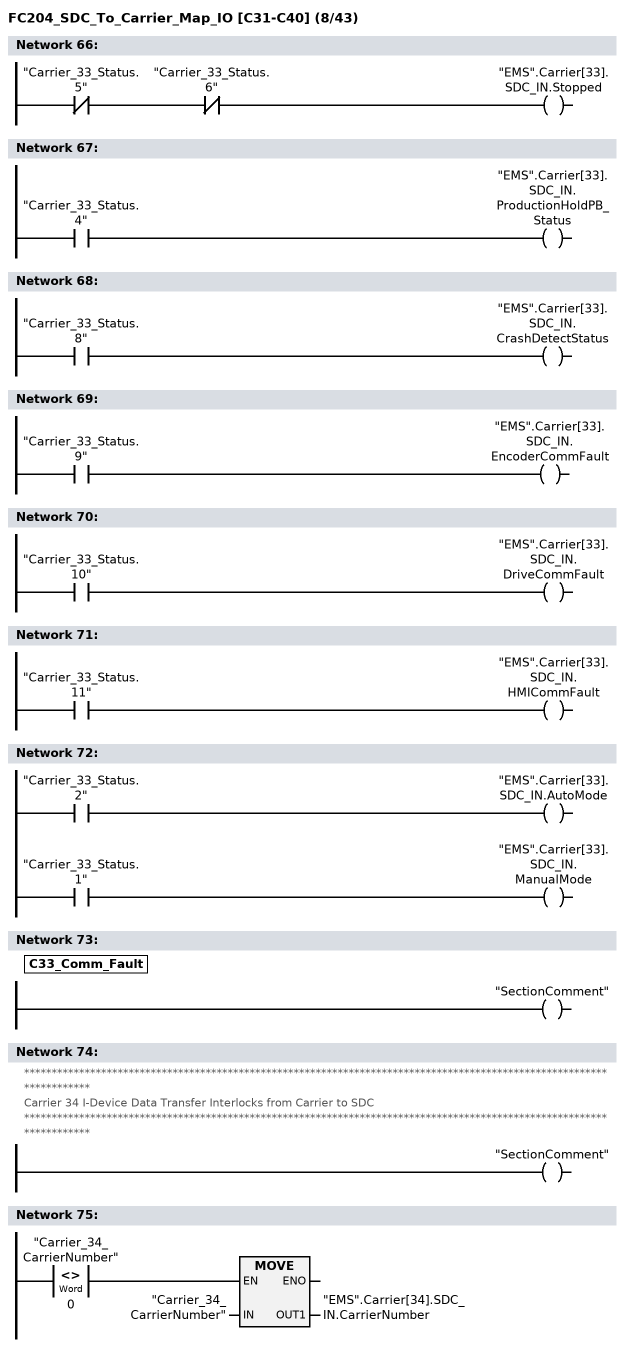
   RUNG wire#powerrail
      I_Contact( "Carrier_33_Status.5" )
      I_Contact( "Carrier_33_Status.6" )
      Coil( "EMS".Carrier[33].SDC_IN.Stopped )
   END_RUNG
   // the same network as SCL:
   "EMS".Carrier[33].SDC_IN.Stopped := NOT "Carrier_33_Status.5" AND NOT "Carrier_33_Status.6";
END_REGION

REGION Network 67
   RUNG wire#powerrail
      Contact( "Carrier_33_Status.4" )
      Coil( "EMS".Carrier[33].SDC_IN.ProductionHoldPB_Status )
   END_RUNG
   // the same network as SCL:
   "EMS".Carrier[33].SDC_IN.ProductionHoldPB_Status := "Carrier_33_Status.4";
END_REGION

REGION Network 68
   RUNG wire#powerrail
      Contact( "Carrier_33_Status.8" )
      Coil( "EMS".Carrier[33].SDC_IN.CrashDetectStatus )
   END_RUNG
   // the same network as SCL:
   "EMS".Carrier[33].SDC_IN.CrashDetectStatus := "Carrier_33_Status.8";
END_REGION

REGION Network 69
   RUNG wire#powerrail
      Contact( "Carrier_33_Status.9" )
      Coil( "EMS".Carrier[33].SDC_IN.EncoderCommFault )
   END_RUNG
   // the same network as SCL:
   "EMS".Carrier[33].SDC_IN.EncoderCommFault := "Carrier_33_Status.9";
END_REGION

REGION Network 70
   RUNG wire#powerrail
      Contact( "Carrier_33_Status.10" )
      Coil( "EMS".Carrier[33].SDC_IN.DriveCommFault )
   END_RUNG
   // the same network as SCL:
   "EMS".Carrier[33].SDC_IN.DriveCommFault := "Carrier_33_Status.10";
END_REGION

REGION Network 71
   RUNG wire#powerrail
      Contact( "Carrier_33_Status.11" )
      Coil( "EMS".Carrier[33].SDC_IN.HMICommFault )
   END_RUNG
   // the same network as SCL:
   "EMS".Carrier[33].SDC_IN.HMICommFault := "Carrier_33_Status.11";
END_REGION

REGION Network 72
   RUNG wire#powerrail
      Contact( "Carrier_33_Status.2" )
      Coil( "EMS".Carrier[33].SDC_IN.AutoMode )
   END_RUNG
   RUNG wire#powerrail
      Contact( "Carrier_33_Status.1" )
      Coil( "EMS".Carrier[33].SDC_IN.ManualMode )
   END_RUNG
   // the same network as SCL:
   "EMS".Carrier[33].SDC_IN.AutoMode := "Carrier_33_Status.2";
   "EMS".Carrier[33].SDC_IN.ManualMode := "Carrier_33_Status.1";
END_REGION

REGION Network 73
   Label( C33_Comm_Fault )
   RUNG wire#powerrail
      Coil( "SectionComment" )
   END_RUNG
   // the same network as SCL:
   C33_Comm_Fault:
   "SectionComment" := TRUE;
END_REGION

REGION Network 74
   // **********************************************************************************************************************
   // 
   // Carrier 34 I-Device Data Transfer Interlocks from Carrier to SDC
   // 
   // **********************************************************************************************************************
   RUNG wire#powerrail
      Coil( "SectionComment" )
   END_RUNG
   // the same network as SCL:
   "SectionComment" := TRUE;
END_REGION

REGION Network 75
   RUNG wire#powerrail
      { S7_Templates := "SrcType := Word" } NE_Contact(in1 := "Carrier_34_CarrierNumber", in2 := 0)
      Move(in := "Carrier_34_CarrierNumber", out1 => "EMS".Carrier[34].SDC_IN.CarrierNumber)
   END_RUNG
   // the same network as SCL:
   IF "Carrier_34_CarrierNumber" <> 0 THEN
       "EMS".Carrier[34].SDC_IN.CarrierNumber := "Carrier_34_CarrierNumber";
   END_IF;
END_REGION

REGION Network 76
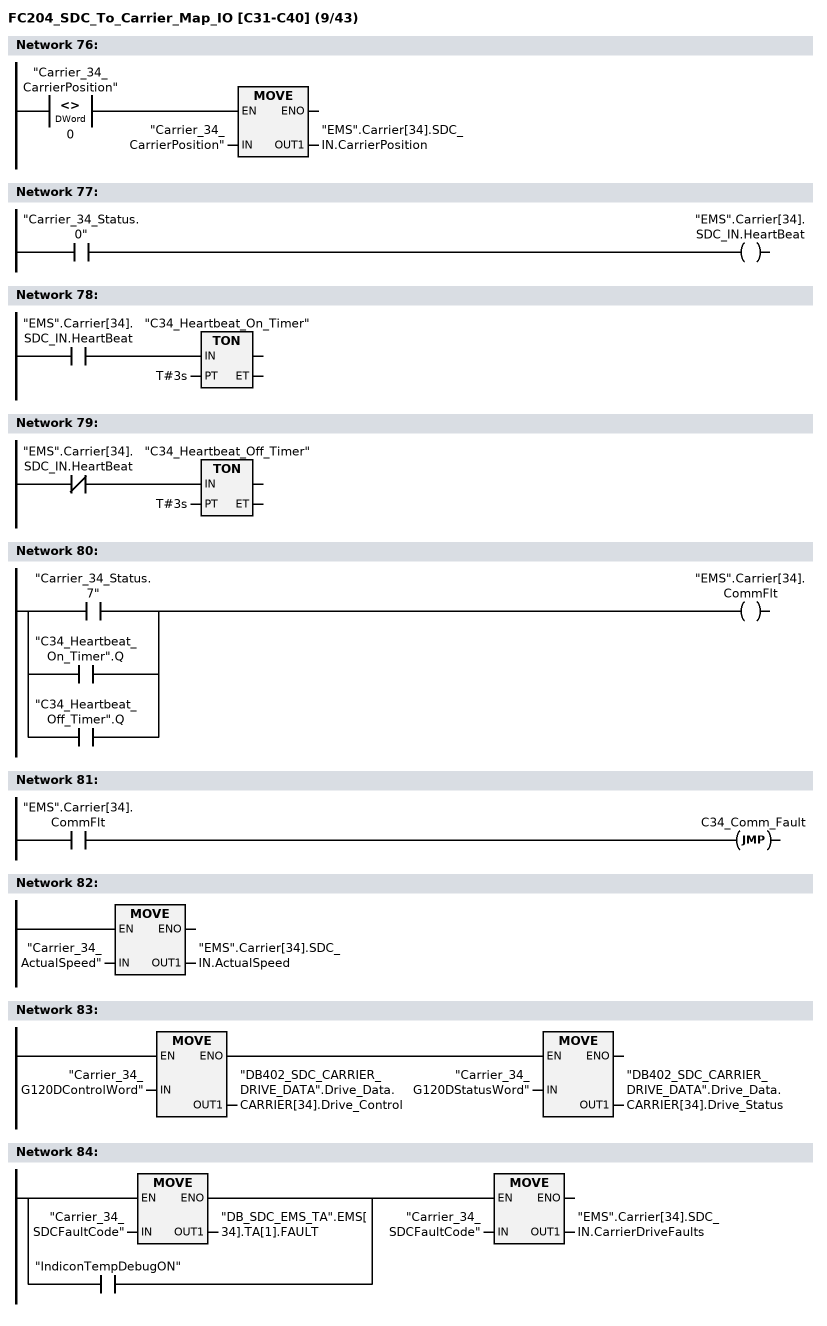
   RUNG wire#powerrail
      { S7_Templates := "SrcType := DWord" } NE_Contact(in1 := "Carrier_34_CarrierPosition", in2 := 0)
      Move(in := "Carrier_34_CarrierPosition", out1 => "EMS".Carrier[34].SDC_IN.CarrierPosition)
   END_RUNG
   // the same network as SCL:
   IF "Carrier_34_CarrierPosition" <> 0 THEN
       "EMS".Carrier[34].SDC_IN.CarrierPosition := "Carrier_34_CarrierPosition";
   END_IF;
END_REGION

REGION Network 77
   RUNG wire#powerrail
      Contact( "Carrier_34_Status.0" )
      Coil( "EMS".Carrier[34].SDC_IN.HeartBeat )
   END_RUNG
   // the same network as SCL:
   "EMS".Carrier[34].SDC_IN.HeartBeat := "Carrier_34_Status.0";
END_REGION

REGION Network 78
   "C34_Heartbeat_On_Timer".TON(IN := "EMS".Carrier[34].SDC_IN.HeartBeat, PT := T#3s);
END_REGION

REGION Network 79
   "C34_Heartbeat_Off_Timer".TON(IN := NOT "EMS".Carrier[34].SDC_IN.HeartBeat, PT := T#3s);
END_REGION

REGION Network 80
   RUNG wire#powerrail
      Contact( "Carrier_34_Status.7" )
      wire#w1
      Coil( "EMS".Carrier[34].CommFlt )
   END_RUNG
   RUNG wire#powerrail
      Contact( "C34_Heartbeat_On_Timer".Q )
   END_RUNG wire#w1
   RUNG wire#powerrail
      Contact( "C34_Heartbeat_Off_Timer".Q )
   END_RUNG wire#w1
   // the same network as SCL:
   "EMS".Carrier[34].CommFlt := "Carrier_34_Status.7" OR "C34_Heartbeat_On_Timer".Q OR "C34_Heartbeat_Off_Timer".Q;
END_REGION

REGION Network 81
   RUNG wire#powerrail
      Contact( "EMS".Carrier[34].CommFlt )
      JumpCoil( C34_Comm_Fault )
   END_RUNG
   // the same network as SCL:
   IF "EMS".Carrier[34].CommFlt THEN GOTO C34_Comm_Fault; END_IF;
END_REGION

REGION Network 82
   RUNG wire#powerrail
      Move(in := "Carrier_34_ActualSpeed", out1 => "EMS".Carrier[34].SDC_IN.ActualSpeed)
   END_RUNG
   // the same network as SCL:
   "EMS".Carrier[34].SDC_IN.ActualSpeed := "Carrier_34_ActualSpeed";
END_REGION

REGION Network 83
   RUNG wire#powerrail
      Move(in := "Carrier_34_G120DControlWord", out1 => "DB402_SDC_CARRIER_DRIVE_DATA".Drive_Data.CARRIER[34].Drive_Control)
      Move(in := "Carrier_34_G120DStatusWord", out1 => "DB402_SDC_CARRIER_DRIVE_DATA".Drive_Data.CARRIER[34].Drive_Status)
   END_RUNG
   // the same network as SCL:
   "DB402_SDC_CARRIER_DRIVE_DATA".Drive_Data.CARRIER[34].Drive_Control := "Carrier_34_G120DControlWord";
   "DB402_SDC_CARRIER_DRIVE_DATA".Drive_Data.CARRIER[34].Drive_Status := "Carrier_34_G120DStatusWord";
END_REGION

REGION Network 84
   RUNG wire#powerrail
      Move(in := "Carrier_34_SDCFaultCode", out1 => "DB_SDC_EMS_TA".EMS[34].TA[1].FAULT)
      wire#w1
      Move(in := "Carrier_34_SDCFaultCode", out1 => "EMS".Carrier[34].SDC_IN.CarrierDriveFaults)
   END_RUNG
   RUNG wire#powerrail
      Contact( "IndiconTempDebugON" )
   END_RUNG wire#w1
   // the same network as SCL:
   "DB_SDC_EMS_TA".EMS[34].TA[1].FAULT := "Carrier_34_SDCFaultCode";
   IF TRUE OR "IndiconTempDebugON" THEN
       "EMS".Carrier[34].SDC_IN.CarrierDriveFaults := "Carrier_34_SDCFaultCode";
   END_IF;
END_REGION

REGION Network 85
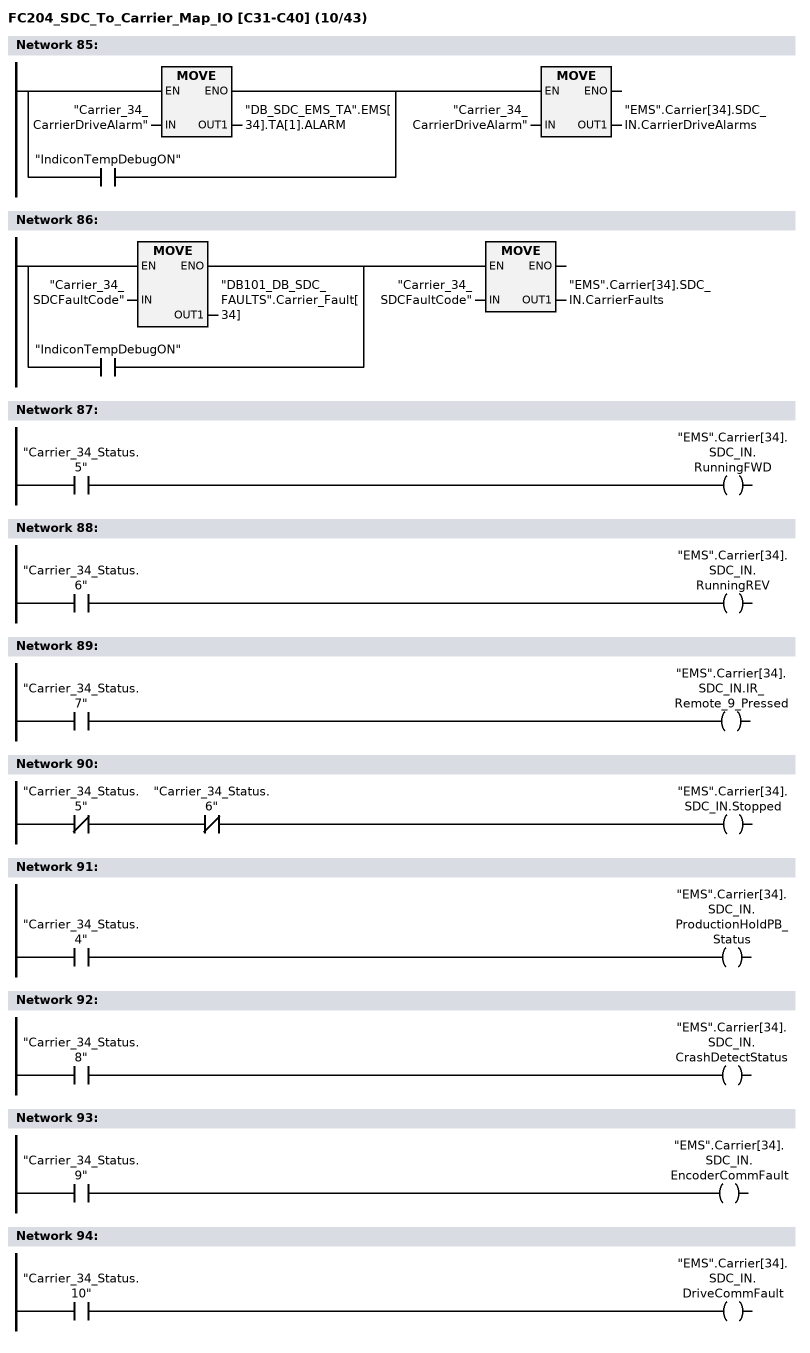
   RUNG wire#powerrail
      Move(in := "Carrier_34_CarrierDriveAlarm", out1 => "DB_SDC_EMS_TA".EMS[34].TA[1].ALARM)
      wire#w1
      Move(in := "Carrier_34_CarrierDriveAlarm", out1 => "EMS".Carrier[34].SDC_IN.CarrierDriveAlarms)
   END_RUNG
   RUNG wire#powerrail
      Contact( "IndiconTempDebugON" )
   END_RUNG wire#w1
   // the same network as SCL:
   "DB_SDC_EMS_TA".EMS[34].TA[1].ALARM := "Carrier_34_CarrierDriveAlarm";
   IF TRUE OR "IndiconTempDebugON" THEN
       "EMS".Carrier[34].SDC_IN.CarrierDriveAlarms := "Carrier_34_CarrierDriveAlarm";
   END_IF;
END_REGION

REGION Network 86
   RUNG wire#powerrail
      Move(in := "Carrier_34_SDCFaultCode", out1 => "DB101_DB_SDC_FAULTS".Carrier_Fault[34])
      wire#w1
      Move(in := "Carrier_34_SDCFaultCode", out1 => "EMS".Carrier[34].SDC_IN.CarrierFaults)
   END_RUNG
   RUNG wire#powerrail
      Contact( "IndiconTempDebugON" )
   END_RUNG wire#w1
   // the same network as SCL:
   "DB101_DB_SDC_FAULTS".Carrier_Fault[34] := "Carrier_34_SDCFaultCode";
   IF TRUE OR "IndiconTempDebugON" THEN
       "EMS".Carrier[34].SDC_IN.CarrierFaults := "Carrier_34_SDCFaultCode";
   END_IF;
END_REGION

REGION Network 87
   RUNG wire#powerrail
      Contact( "Carrier_34_Status.5" )
      Coil( "EMS".Carrier[34].SDC_IN.RunningFWD )
   END_RUNG
   // the same network as SCL:
   "EMS".Carrier[34].SDC_IN.RunningFWD := "Carrier_34_Status.5";
END_REGION

REGION Network 88
   RUNG wire#powerrail
      Contact( "Carrier_34_Status.6" )
      Coil( "EMS".Carrier[34].SDC_IN.RunningREV )
   END_RUNG
   // the same network as SCL:
   "EMS".Carrier[34].SDC_IN.RunningREV := "Carrier_34_Status.6";
END_REGION

REGION Network 89
   RUNG wire#powerrail
      Contact( "Carrier_34_Status.7" )
      Coil( "EMS".Carrier[34].SDC_IN.IR_Remote_9_Pressed )
   END_RUNG
   // the same network as SCL:
   "EMS".Carrier[34].SDC_IN.IR_Remote_9_Pressed := "Carrier_34_Status.7";
END_REGION

REGION Network 90
   RUNG wire#powerrail
      I_Contact( "Carrier_34_Status.5" )
      I_Contact( "Carrier_34_Status.6" )
      Coil( "EMS".Carrier[34].SDC_IN.Stopped )
   END_RUNG
   // the same network as SCL:
   "EMS".Carrier[34].SDC_IN.Stopped := NOT "Carrier_34_Status.5" AND NOT "Carrier_34_Status.6";
END_REGION

REGION Network 91
   RUNG wire#powerrail
      Contact( "Carrier_34_Status.4" )
      Coil( "EMS".Carrier[34].SDC_IN.ProductionHoldPB_Status )
   END_RUNG
   // the same network as SCL:
   "EMS".Carrier[34].SDC_IN.ProductionHoldPB_Status := "Carrier_34_Status.4";
END_REGION

REGION Network 92
   RUNG wire#powerrail
      Contact( "Carrier_34_Status.8" )
      Coil( "EMS".Carrier[34].SDC_IN.CrashDetectStatus )
   END_RUNG
   // the same network as SCL:
   "EMS".Carrier[34].SDC_IN.CrashDetectStatus := "Carrier_34_Status.8";
END_REGION

REGION Network 93
   RUNG wire#powerrail
      Contact( "Carrier_34_Status.9" )
      Coil( "EMS".Carrier[34].SDC_IN.EncoderCommFault )
   END_RUNG
   // the same network as SCL:
   "EMS".Carrier[34].SDC_IN.EncoderCommFault := "Carrier_34_Status.9";
END_REGION

REGION Network 94
   RUNG wire#powerrail
      Contact( "Carrier_34_Status.10" )
      Coil( "EMS".Carrier[34].SDC_IN.DriveCommFault )
   END_RUNG
   // the same network as SCL:
   "EMS".Carrier[34].SDC_IN.DriveCommFault := "Carrier_34_Status.10";
END_REGION

REGION Network 95
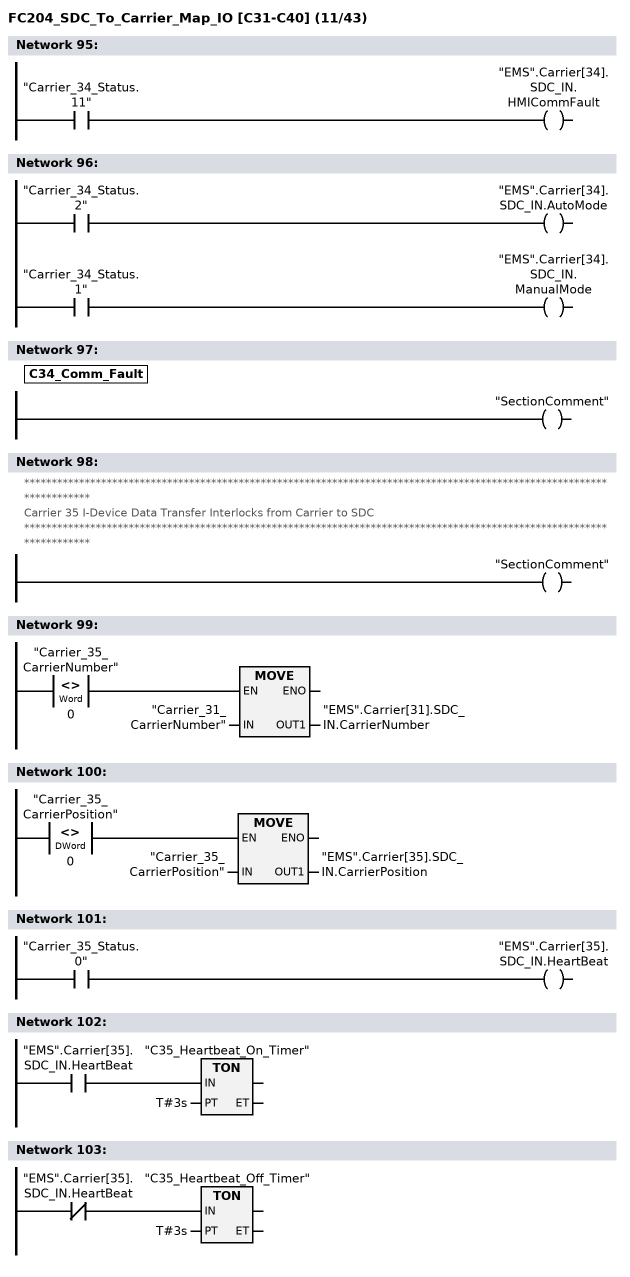
   RUNG wire#powerrail
      Contact( "Carrier_34_Status.11" )
      Coil( "EMS".Carrier[34].SDC_IN.HMICommFault )
   END_RUNG
   // the same network as SCL:
   "EMS".Carrier[34].SDC_IN.HMICommFault := "Carrier_34_Status.11";
END_REGION

REGION Network 96
   RUNG wire#powerrail
      Contact( "Carrier_34_Status.2" )
      Coil( "EMS".Carrier[34].SDC_IN.AutoMode )
   END_RUNG
   RUNG wire#powerrail
      Contact( "Carrier_34_Status.1" )
      Coil( "EMS".Carrier[34].SDC_IN.ManualMode )
   END_RUNG
   // the same network as SCL:
   "EMS".Carrier[34].SDC_IN.AutoMode := "Carrier_34_Status.2";
   "EMS".Carrier[34].SDC_IN.ManualMode := "Carrier_34_Status.1";
END_REGION

REGION Network 97
   Label( C34_Comm_Fault )
   RUNG wire#powerrail
      Coil( "SectionComment" )
   END_RUNG
   // the same network as SCL:
   C34_Comm_Fault:
   "SectionComment" := TRUE;
END_REGION

REGION Network 98
   // **********************************************************************************************************************
   // 
   // Carrier 35 I-Device Data Transfer Interlocks from Carrier to SDC
   // 
   // **********************************************************************************************************************
   RUNG wire#powerrail
      Coil( "SectionComment" )
   END_RUNG
   // the same network as SCL:
   "SectionComment" := TRUE;
END_REGION

REGION Network 99
   RUNG wire#powerrail
      { S7_Templates := "SrcType := Word" } NE_Contact(in1 := "Carrier_35_CarrierNumber", in2 := 0)
      Move(in := "Carrier_31_CarrierNumber", out1 => "EMS".Carrier[31].SDC_IN.CarrierNumber)
   END_RUNG
   // the same network as SCL:
   IF "Carrier_35_CarrierNumber" <> 0 THEN
       "EMS".Carrier[31].SDC_IN.CarrierNumber := "Carrier_31_CarrierNumber";
   END_IF;
END_REGION

REGION Network 100
   RUNG wire#powerrail
      { S7_Templates := "SrcType := DWord" } NE_Contact(in1 := "Carrier_35_CarrierPosition", in2 := 0)
      Move(in := "Carrier_35_CarrierPosition", out1 => "EMS".Carrier[35].SDC_IN.CarrierPosition)
   END_RUNG
   // the same network as SCL:
   IF "Carrier_35_CarrierPosition" <> 0 THEN
       "EMS".Carrier[35].SDC_IN.CarrierPosition := "Carrier_35_CarrierPosition";
   END_IF;
END_REGION

REGION Network 101
   RUNG wire#powerrail
      Contact( "Carrier_35_Status.0" )
      Coil( "EMS".Carrier[35].SDC_IN.HeartBeat )
   END_RUNG
   // the same network as SCL:
   "EMS".Carrier[35].SDC_IN.HeartBeat := "Carrier_35_Status.0";
END_REGION

REGION Network 102
   "C35_Heartbeat_On_Timer".TON(IN := "EMS".Carrier[35].SDC_IN.HeartBeat, PT := T#3s);
END_REGION

REGION Network 103
   "C35_Heartbeat_Off_Timer".TON(IN := NOT "EMS".Carrier[35].SDC_IN.HeartBeat, PT := T#3s);
END_REGION

REGION Network 104
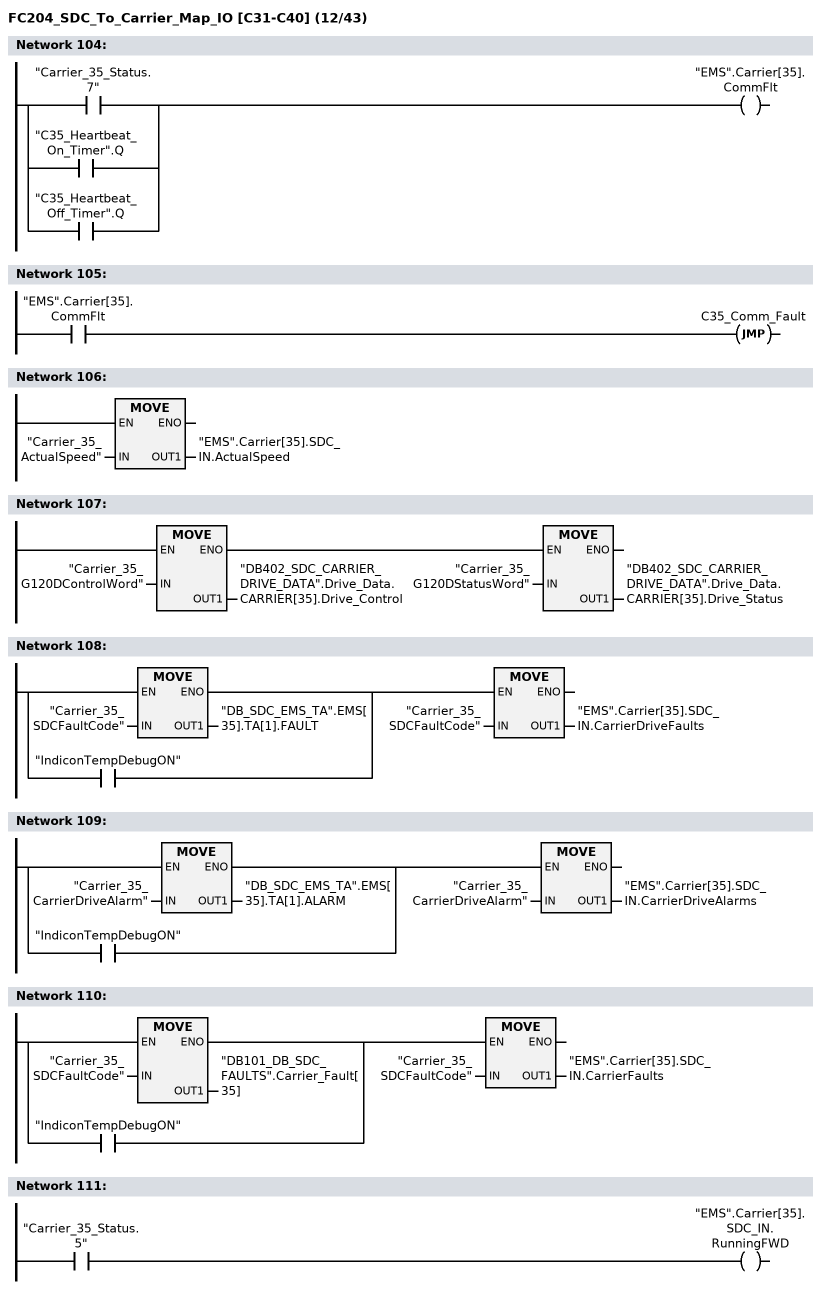
   RUNG wire#powerrail
      Contact( "Carrier_35_Status.7" )
      wire#w1
      Coil( "EMS".Carrier[35].CommFlt )
   END_RUNG
   RUNG wire#powerrail
      Contact( "C35_Heartbeat_On_Timer".Q )
   END_RUNG wire#w1
   RUNG wire#powerrail
      Contact( "C35_Heartbeat_Off_Timer".Q )
   END_RUNG wire#w1
   // the same network as SCL:
   "EMS".Carrier[35].CommFlt := "Carrier_35_Status.7" OR "C35_Heartbeat_On_Timer".Q OR "C35_Heartbeat_Off_Timer".Q;
END_REGION

REGION Network 105
   RUNG wire#powerrail
      Contact( "EMS".Carrier[35].CommFlt )
      JumpCoil( C35_Comm_Fault )
   END_RUNG
   // the same network as SCL:
   IF "EMS".Carrier[35].CommFlt THEN GOTO C35_Comm_Fault; END_IF;
END_REGION

REGION Network 106
   RUNG wire#powerrail
      Move(in := "Carrier_35_ActualSpeed", out1 => "EMS".Carrier[35].SDC_IN.ActualSpeed)
   END_RUNG
   // the same network as SCL:
   "EMS".Carrier[35].SDC_IN.ActualSpeed := "Carrier_35_ActualSpeed";
END_REGION

REGION Network 107
   RUNG wire#powerrail
      Move(in := "Carrier_35_G120DControlWord", out1 => "DB402_SDC_CARRIER_DRIVE_DATA".Drive_Data.CARRIER[35].Drive_Control)
      Move(in := "Carrier_35_G120DStatusWord", out1 => "DB402_SDC_CARRIER_DRIVE_DATA".Drive_Data.CARRIER[35].Drive_Status)
   END_RUNG
   // the same network as SCL:
   "DB402_SDC_CARRIER_DRIVE_DATA".Drive_Data.CARRIER[35].Drive_Control := "Carrier_35_G120DControlWord";
   "DB402_SDC_CARRIER_DRIVE_DATA".Drive_Data.CARRIER[35].Drive_Status := "Carrier_35_G120DStatusWord";
END_REGION

REGION Network 108
   RUNG wire#powerrail
      Move(in := "Carrier_35_SDCFaultCode", out1 => "DB_SDC_EMS_TA".EMS[35].TA[1].FAULT)
      wire#w1
      Move(in := "Carrier_35_SDCFaultCode", out1 => "EMS".Carrier[35].SDC_IN.CarrierDriveFaults)
   END_RUNG
   RUNG wire#powerrail
      Contact( "IndiconTempDebugON" )
   END_RUNG wire#w1
   // the same network as SCL:
   "DB_SDC_EMS_TA".EMS[35].TA[1].FAULT := "Carrier_35_SDCFaultCode";
   IF TRUE OR "IndiconTempDebugON" THEN
       "EMS".Carrier[35].SDC_IN.CarrierDriveFaults := "Carrier_35_SDCFaultCode";
   END_IF;
END_REGION

REGION Network 109
   RUNG wire#powerrail
      Move(in := "Carrier_35_CarrierDriveAlarm", out1 => "DB_SDC_EMS_TA".EMS[35].TA[1].ALARM)
      wire#w1
      Move(in := "Carrier_35_CarrierDriveAlarm", out1 => "EMS".Carrier[35].SDC_IN.CarrierDriveAlarms)
   END_RUNG
   RUNG wire#powerrail
      Contact( "IndiconTempDebugON" )
   END_RUNG wire#w1
   // the same network as SCL:
   "DB_SDC_EMS_TA".EMS[35].TA[1].ALARM := "Carrier_35_CarrierDriveAlarm";
   IF TRUE OR "IndiconTempDebugON" THEN
       "EMS".Carrier[35].SDC_IN.CarrierDriveAlarms := "Carrier_35_CarrierDriveAlarm";
   END_IF;
END_REGION

REGION Network 110
   RUNG wire#powerrail
      Move(in := "Carrier_35_SDCFaultCode", out1 => "DB101_DB_SDC_FAULTS".Carrier_Fault[35])
      wire#w1
      Move(in := "Carrier_35_SDCFaultCode", out1 => "EMS".Carrier[35].SDC_IN.CarrierFaults)
   END_RUNG
   RUNG wire#powerrail
      Contact( "IndiconTempDebugON" )
   END_RUNG wire#w1
   // the same network as SCL:
   "DB101_DB_SDC_FAULTS".Carrier_Fault[35] := "Carrier_35_SDCFaultCode";
   IF TRUE OR "IndiconTempDebugON" THEN
       "EMS".Carrier[35].SDC_IN.CarrierFaults := "Carrier_35_SDCFaultCode";
   END_IF;
END_REGION

REGION Network 111
   RUNG wire#powerrail
      Contact( "Carrier_35_Status.5" )
      Coil( "EMS".Carrier[35].SDC_IN.RunningFWD )
   END_RUNG
   // the same network as SCL:
   "EMS".Carrier[35].SDC_IN.RunningFWD := "Carrier_35_Status.5";
END_REGION

REGION Network 112
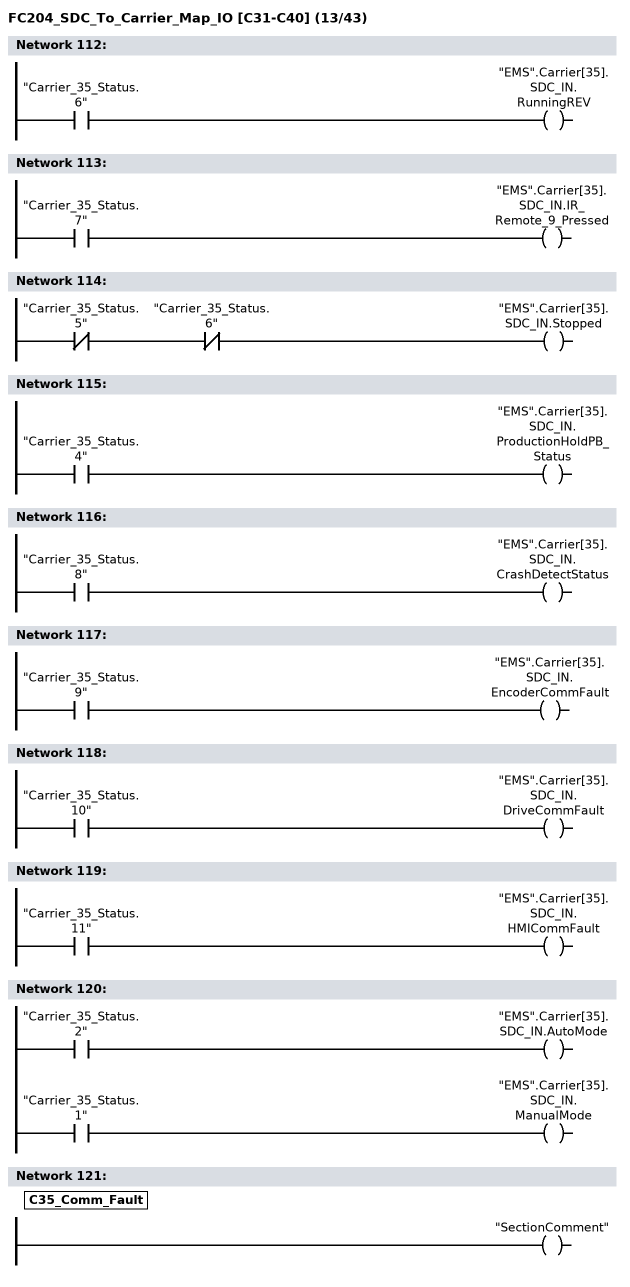
   RUNG wire#powerrail
      Contact( "Carrier_35_Status.6" )
      Coil( "EMS".Carrier[35].SDC_IN.RunningREV )
   END_RUNG
   // the same network as SCL:
   "EMS".Carrier[35].SDC_IN.RunningREV := "Carrier_35_Status.6";
END_REGION

REGION Network 113
   RUNG wire#powerrail
      Contact( "Carrier_35_Status.7" )
      Coil( "EMS".Carrier[35].SDC_IN.IR_Remote_9_Pressed )
   END_RUNG
   // the same network as SCL:
   "EMS".Carrier[35].SDC_IN.IR_Remote_9_Pressed := "Carrier_35_Status.7";
END_REGION

REGION Network 114
   RUNG wire#powerrail
      I_Contact( "Carrier_35_Status.5" )
      I_Contact( "Carrier_35_Status.6" )
      Coil( "EMS".Carrier[35].SDC_IN.Stopped )
   END_RUNG
   // the same network as SCL:
   "EMS".Carrier[35].SDC_IN.Stopped := NOT "Carrier_35_Status.5" AND NOT "Carrier_35_Status.6";
END_REGION

REGION Network 115
   RUNG wire#powerrail
      Contact( "Carrier_35_Status.4" )
      Coil( "EMS".Carrier[35].SDC_IN.ProductionHoldPB_Status )
   END_RUNG
   // the same network as SCL:
   "EMS".Carrier[35].SDC_IN.ProductionHoldPB_Status := "Carrier_35_Status.4";
END_REGION

REGION Network 116
   RUNG wire#powerrail
      Contact( "Carrier_35_Status.8" )
      Coil( "EMS".Carrier[35].SDC_IN.CrashDetectStatus )
   END_RUNG
   // the same network as SCL:
   "EMS".Carrier[35].SDC_IN.CrashDetectStatus := "Carrier_35_Status.8";
END_REGION

REGION Network 117
   RUNG wire#powerrail
      Contact( "Carrier_35_Status.9" )
      Coil( "EMS".Carrier[35].SDC_IN.EncoderCommFault )
   END_RUNG
   // the same network as SCL:
   "EMS".Carrier[35].SDC_IN.EncoderCommFault := "Carrier_35_Status.9";
END_REGION

REGION Network 118
   RUNG wire#powerrail
      Contact( "Carrier_35_Status.10" )
      Coil( "EMS".Carrier[35].SDC_IN.DriveCommFault )
   END_RUNG
   // the same network as SCL:
   "EMS".Carrier[35].SDC_IN.DriveCommFault := "Carrier_35_Status.10";
END_REGION

REGION Network 119
   RUNG wire#powerrail
      Contact( "Carrier_35_Status.11" )
      Coil( "EMS".Carrier[35].SDC_IN.HMICommFault )
   END_RUNG
   // the same network as SCL:
   "EMS".Carrier[35].SDC_IN.HMICommFault := "Carrier_35_Status.11";
END_REGION

REGION Network 120
   RUNG wire#powerrail
      Contact( "Carrier_35_Status.2" )
      Coil( "EMS".Carrier[35].SDC_IN.AutoMode )
   END_RUNG
   RUNG wire#powerrail
      Contact( "Carrier_35_Status.1" )
      Coil( "EMS".Carrier[35].SDC_IN.ManualMode )
   END_RUNG
   // the same network as SCL:
   "EMS".Carrier[35].SDC_IN.AutoMode := "Carrier_35_Status.2";
   "EMS".Carrier[35].SDC_IN.ManualMode := "Carrier_35_Status.1";
END_REGION

REGION Network 121
   Label( C35_Comm_Fault )
   RUNG wire#powerrail
      Coil( "SectionComment" )
   END_RUNG
   // the same network as SCL:
   C35_Comm_Fault:
   "SectionComment" := TRUE;
END_REGION

REGION Network 122
   // **********************************************************************************************************************
   // 
   // Carrier 36 I-Device Data Transfer Interlocks from Carrier to SDC
   // 
   // **********************************************************************************************************************
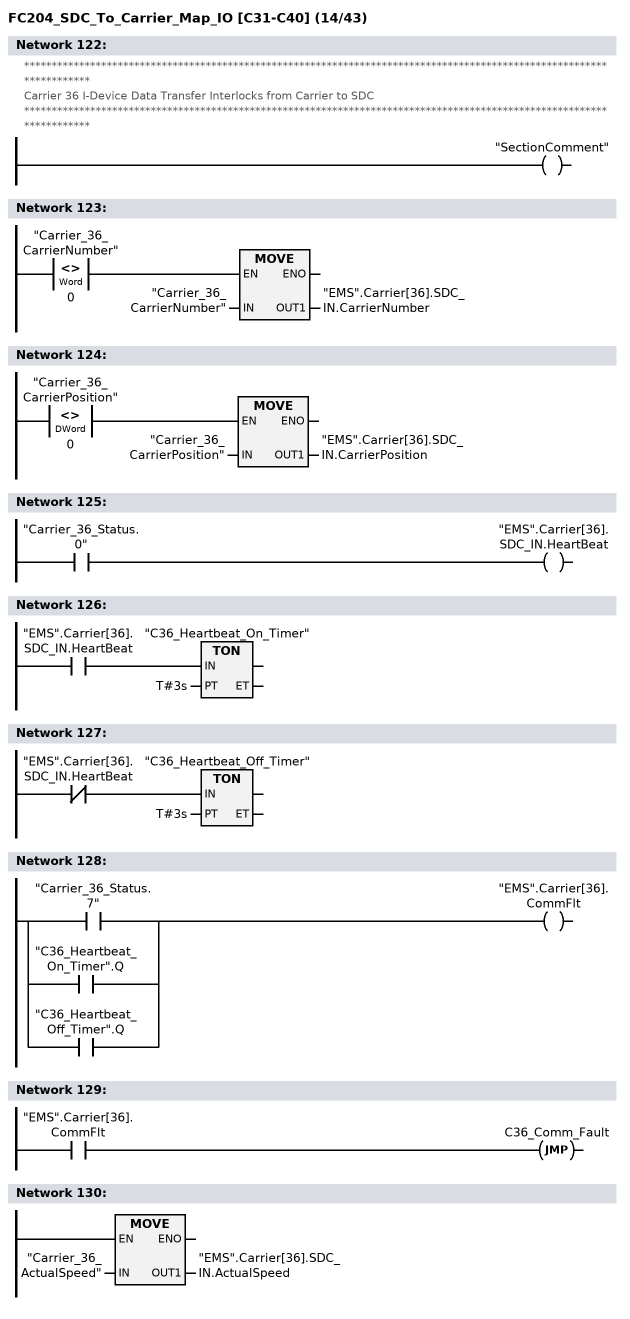
   RUNG wire#powerrail
      Coil( "SectionComment" )
   END_RUNG
   // the same network as SCL:
   "SectionComment" := TRUE;
END_REGION

REGION Network 123
   RUNG wire#powerrail
      { S7_Templates := "SrcType := Word" } NE_Contact(in1 := "Carrier_36_CarrierNumber", in2 := 0)
      Move(in := "Carrier_36_CarrierNumber", out1 => "EMS".Carrier[36].SDC_IN.CarrierNumber)
   END_RUNG
   // the same network as SCL:
   IF "Carrier_36_CarrierNumber" <> 0 THEN
       "EMS".Carrier[36].SDC_IN.CarrierNumber := "Carrier_36_CarrierNumber";
   END_IF;
END_REGION

REGION Network 124
   RUNG wire#powerrail
      { S7_Templates := "SrcType := DWord" } NE_Contact(in1 := "Carrier_36_CarrierPosition", in2 := 0)
      Move(in := "Carrier_36_CarrierPosition", out1 => "EMS".Carrier[36].SDC_IN.CarrierPosition)
   END_RUNG
   // the same network as SCL:
   IF "Carrier_36_CarrierPosition" <> 0 THEN
       "EMS".Carrier[36].SDC_IN.CarrierPosition := "Carrier_36_CarrierPosition";
   END_IF;
END_REGION

REGION Network 125
   RUNG wire#powerrail
      Contact( "Carrier_36_Status.0" )
      Coil( "EMS".Carrier[36].SDC_IN.HeartBeat )
   END_RUNG
   // the same network as SCL:
   "EMS".Carrier[36].SDC_IN.HeartBeat := "Carrier_36_Status.0";
END_REGION

REGION Network 126
   "C36_Heartbeat_On_Timer".TON(IN := "EMS".Carrier[36].SDC_IN.HeartBeat, PT := T#3s);
END_REGION

REGION Network 127
   "C36_Heartbeat_Off_Timer".TON(IN := NOT "EMS".Carrier[36].SDC_IN.HeartBeat, PT := T#3s);
END_REGION

REGION Network 128
   RUNG wire#powerrail
      Contact( "Carrier_36_Status.7" )
      wire#w1
      Coil( "EMS".Carrier[36].CommFlt )
   END_RUNG
   RUNG wire#powerrail
      Contact( "C36_Heartbeat_On_Timer".Q )
   END_RUNG wire#w1
   RUNG wire#powerrail
      Contact( "C36_Heartbeat_Off_Timer".Q )
   END_RUNG wire#w1
   // the same network as SCL:
   "EMS".Carrier[36].CommFlt := "Carrier_36_Status.7" OR "C36_Heartbeat_On_Timer".Q OR "C36_Heartbeat_Off_Timer".Q;
END_REGION

REGION Network 129
   RUNG wire#powerrail
      Contact( "EMS".Carrier[36].CommFlt )
      JumpCoil( C36_Comm_Fault )
   END_RUNG
   // the same network as SCL:
   IF "EMS".Carrier[36].CommFlt THEN GOTO C36_Comm_Fault; END_IF;
END_REGION

REGION Network 130
   RUNG wire#powerrail
      Move(in := "Carrier_36_ActualSpeed", out1 => "EMS".Carrier[36].SDC_IN.ActualSpeed)
   END_RUNG
   // the same network as SCL:
   "EMS".Carrier[36].SDC_IN.ActualSpeed := "Carrier_36_ActualSpeed";
END_REGION

REGION Network 131
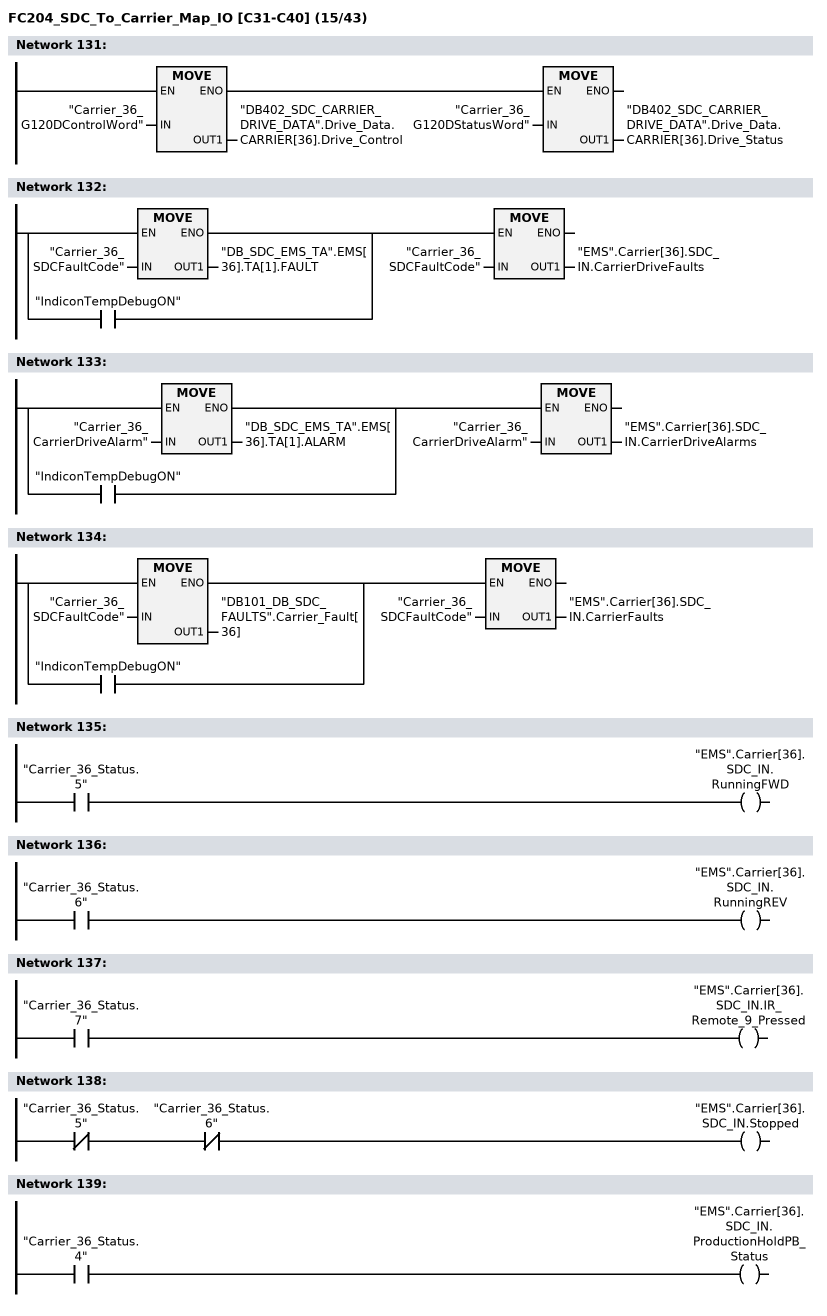
   RUNG wire#powerrail
      Move(in := "Carrier_36_G120DControlWord", out1 => "DB402_SDC_CARRIER_DRIVE_DATA".Drive_Data.CARRIER[36].Drive_Control)
      Move(in := "Carrier_36_G120DStatusWord", out1 => "DB402_SDC_CARRIER_DRIVE_DATA".Drive_Data.CARRIER[36].Drive_Status)
   END_RUNG
   // the same network as SCL:
   "DB402_SDC_CARRIER_DRIVE_DATA".Drive_Data.CARRIER[36].Drive_Control := "Carrier_36_G120DControlWord";
   "DB402_SDC_CARRIER_DRIVE_DATA".Drive_Data.CARRIER[36].Drive_Status := "Carrier_36_G120DStatusWord";
END_REGION

REGION Network 132
   RUNG wire#powerrail
      Move(in := "Carrier_36_SDCFaultCode", out1 => "DB_SDC_EMS_TA".EMS[36].TA[1].FAULT)
      wire#w1
      Move(in := "Carrier_36_SDCFaultCode", out1 => "EMS".Carrier[36].SDC_IN.CarrierDriveFaults)
   END_RUNG
   RUNG wire#powerrail
      Contact( "IndiconTempDebugON" )
   END_RUNG wire#w1
   // the same network as SCL:
   "DB_SDC_EMS_TA".EMS[36].TA[1].FAULT := "Carrier_36_SDCFaultCode";
   IF TRUE OR "IndiconTempDebugON" THEN
       "EMS".Carrier[36].SDC_IN.CarrierDriveFaults := "Carrier_36_SDCFaultCode";
   END_IF;
END_REGION

REGION Network 133
   RUNG wire#powerrail
      Move(in := "Carrier_36_CarrierDriveAlarm", out1 => "DB_SDC_EMS_TA".EMS[36].TA[1].ALARM)
      wire#w1
      Move(in := "Carrier_36_CarrierDriveAlarm", out1 => "EMS".Carrier[36].SDC_IN.CarrierDriveAlarms)
   END_RUNG
   RUNG wire#powerrail
      Contact( "IndiconTempDebugON" )
   END_RUNG wire#w1
   // the same network as SCL:
   "DB_SDC_EMS_TA".EMS[36].TA[1].ALARM := "Carrier_36_CarrierDriveAlarm";
   IF TRUE OR "IndiconTempDebugON" THEN
       "EMS".Carrier[36].SDC_IN.CarrierDriveAlarms := "Carrier_36_CarrierDriveAlarm";
   END_IF;
END_REGION

REGION Network 134
   RUNG wire#powerrail
      Move(in := "Carrier_36_SDCFaultCode", out1 => "DB101_DB_SDC_FAULTS".Carrier_Fault[36])
      wire#w1
      Move(in := "Carrier_36_SDCFaultCode", out1 => "EMS".Carrier[36].SDC_IN.CarrierFaults)
   END_RUNG
   RUNG wire#powerrail
      Contact( "IndiconTempDebugON" )
   END_RUNG wire#w1
   // the same network as SCL:
   "DB101_DB_SDC_FAULTS".Carrier_Fault[36] := "Carrier_36_SDCFaultCode";
   IF TRUE OR "IndiconTempDebugON" THEN
       "EMS".Carrier[36].SDC_IN.CarrierFaults := "Carrier_36_SDCFaultCode";
   END_IF;
END_REGION

REGION Network 135
   RUNG wire#powerrail
      Contact( "Carrier_36_Status.5" )
      Coil( "EMS".Carrier[36].SDC_IN.RunningFWD )
   END_RUNG
   // the same network as SCL:
   "EMS".Carrier[36].SDC_IN.RunningFWD := "Carrier_36_Status.5";
END_REGION

REGION Network 136
   RUNG wire#powerrail
      Contact( "Carrier_36_Status.6" )
      Coil( "EMS".Carrier[36].SDC_IN.RunningREV )
   END_RUNG
   // the same network as SCL:
   "EMS".Carrier[36].SDC_IN.RunningREV := "Carrier_36_Status.6";
END_REGION

REGION Network 137
   RUNG wire#powerrail
      Contact( "Carrier_36_Status.7" )
      Coil( "EMS".Carrier[36].SDC_IN.IR_Remote_9_Pressed )
   END_RUNG
   // the same network as SCL:
   "EMS".Carrier[36].SDC_IN.IR_Remote_9_Pressed := "Carrier_36_Status.7";
END_REGION

REGION Network 138
   RUNG wire#powerrail
      I_Contact( "Carrier_36_Status.5" )
      I_Contact( "Carrier_36_Status.6" )
      Coil( "EMS".Carrier[36].SDC_IN.Stopped )
   END_RUNG
   // the same network as SCL:
   "EMS".Carrier[36].SDC_IN.Stopped := NOT "Carrier_36_Status.5" AND NOT "Carrier_36_Status.6";
END_REGION

REGION Network 139
   RUNG wire#powerrail
      Contact( "Carrier_36_Status.4" )
      Coil( "EMS".Carrier[36].SDC_IN.ProductionHoldPB_Status )
   END_RUNG
   // the same network as SCL:
   "EMS".Carrier[36].SDC_IN.ProductionHoldPB_Status := "Carrier_36_Status.4";
END_REGION

REGION Network 140
